   		UOWHF_Result[0].31:=0;
   		UOWHF_Result[1]:=UOWHF_Result[1] + 783475357+UOWHF_Add_c;
   		UOWHF_Add_c.1:=UOWHF_Result[1].31;
   		UOWHF_Result[1].31:=0;
   		UOWHF_Result[2]:=UOWHF_Result[2] + 293797280+UOWHF_Add_c;
   		UOWHF_Add_c.2:=UOWHF_Result[2].31;
   		UOWHF_Result[2].31:=0;
   		UOWHF_Result[3]:=UOWHF_Result[3] + 185650386+UOWHF_Add_c;
   		UOWHF_Add_c.3:=UOWHF_Result[3].31;
   		UOWHF_Result[3].31:=0;
   		UOWHF_Result[4]:=UOWHF_Result[4] + 976456778+UOWHF_Add_c;
   		UOWHF_Add_c.4:=UOWHF_Result[4].31;
   		UOWHF_Result[4].31:=0;
   		UOWHF_Result[5]:=UOWHF_Result[5] + 1830429797+UOWHF_Add_c;
   		UOWHF_Add_c.5:=UOWHF_Result[5].31;
   		UOWHF_Result[5].31:=0;
   		UOWHF_Result[6]:=UOWHF_Result[6] + 346921929+UOWHF_Add_c;
   		UOWHF_Add_c.6:=UOWHF_Result[6].31;
   		UOWHF_Result[6].31:=0;
   	End_If;
   	If UOWHF_Msg[1].[3] Then
   		UOWHF_Result[0]:=UOWHF_Result[0] + 542356735+UOWHF_Add_c;
   		UOWHF_Add_c.0:=UOWHF_Result[0].31;
   		UOWHF_Result[0].31:=0;
   		UOWHF_Result[1]:=UOWHF_Result[1] + 1471465957+UOWHF_Add_c;
   		UOWHF_Add_c.1:=UOWHF_Result[1].31;
   		UOWHF_Result[1].31:=0;
   		UOWHF_Result[2]:=UOWHF_Result[2] + 880885546+UOWHF_Add_c;
   		UOWHF_Add_c.2:=UOWHF_Result[2].31;
   		UOWHF_Result[2].31:=0;
   		UOWHF_Result[3]:=UOWHF_Result[3] + 1420715233+UOWHF_Add_c;
   		UOWHF_Add_c.3:=UOWHF_Result[3].31;
   		UOWHF_Result[3].31:=0;
   		UOWHF_Result[4]:=UOWHF_Result[4] + 974859291+UOWHF_Add_c;
   		UOWHF_Add_c.4:=UOWHF_Result[4].31;
   		UOWHF_Result[4].31:=0;
   		UOWHF_Result[5]:=UOWHF_Result[5] + 2135033399+UOWHF_Add_c;
   		UOWHF_Add_c.5:=UOWHF_Result[5].31;
   		UOWHF_Result[5].31:=0;
   		UOWHF_Result[6]:=UOWHF_Result[6] + 991907939+UOWHF_Add_c;
   		UOWHF_Add_c.6:=UOWHF_Result[6].31;
   		UOWHF_Result[6].31:=0;
   	End_If;
   	If UOWHF_Msg[1].[4] Then
   		UOWHF_Result[0]:=UOWHF_Result[0] + 233841843+UOWHF_Add_c;
   		UOWHF_Add_c.0:=UOWHF_Result[0].31;
   		UOWHF_Result[0].31:=0;
   		UOWHF_Result[1]:=UOWHF_Result[1] + 422275350+UOWHF_Add_c;
   		UOWHF_Add_c.1:=UOWHF_Result[1].31;
   		UOWHF_Result[1].31:=0;
   		UOWHF_Result[2]:=UOWHF_Result[2] + 758599260+UOWHF_Add_c;
   		UOWHF_Add_c.2:=UOWHF_Result[2].31;
   		UOWHF_Result[2].31:=0;
   		UOWHF_Result[3]:=UOWHF_Result[3] + 1065130774+UOWHF_Add_c;
   		UOWHF_Add_c.3:=UOWHF_Result[3].31;
   		UOWHF_Result[3].31:=0;
   		UOWHF_Result[4]:=UOWHF_Result[4] + 2001915225+UOWHF_Add_c;
   		UOWHF_Add_c.4:=UOWHF_Result[4].31;
   		UOWHF_Result[4].31:=0;
   		UOWHF_Result[5]:=UOWHF_Result[5] + 545495531+UOWHF_Add_c;
   		UOWHF_Add_c.5:=UOWHF_Result[5].31;
   		UOWHF_Result[5].31:=0;
   		UOWHF_Result[6]:=UOWHF_Result[6] + 296068018+UOWHF_Add_c;
   		UOWHF_Add_c.6:=UOWHF_Result[6].31;
   		UOWHF_Result[6].31:=0;
   	End_If;
   	If UOWHF_Msg[1].[5] Then
   		UOWHF_Result[0]:=UOWHF_Result[0] + 5724122+UOWHF_Add_c;
   		UOWHF_Add_c.0:=UOWHF_Result[0].31;
   		UOWHF_Result[0].31:=0;
   		UOWHF_Result[1]:=UOWHF_Result[1] + 218649241+UOWHF_Add_c;
   		UOWHF_Add_c.1:=UOWHF_Result[1].31;
   		UOWHF_Result[1].31:=0;
   		UOWHF_Result[2]:=UOWHF_Result[2] + 238121106+UOWHF_Add_c;
   		UOWHF_Add_c.2:=UOWHF_Result[2].31;
   		UOWHF_Result[2].31:=0;
   		UOWHF_Result[3]:=UOWHF_Result[3] + 729241869+UOWHF_Add_c;
   		UOWHF_Add_c.3:=UOWHF_Result[3].31;
   		UOWHF_Result[3].31:=0;
   		UOWHF_Result[4]:=UOWHF_Result[4] + 1651167024+UOWHF_Add_c;
   		UOWHF_Add_c.4:=UOWHF_Result[4].31;
   		UOWHF_Result[4].31:=0;
   		UOWHF_Result[5]:=UOWHF_Result[5] + 2110643339+UOWHF_Add_c;
   		UOWHF_Add_c.5:=UOWHF_Result[5].31;
   		UOWHF_Result[5].31:=0;
   		UOWHF_Result[6]:=UOWHF_Result[6] + 1917524854+UOWHF_Add_c;
   		UOWHF_Add_c.6:=UOWHF_Result[6].31;
   		UOWHF_Result[6].31:=0;
   	End_If;
   	If UOWHF_Msg[1].[6] Then
   		UOWHF_Result[0]:=UOWHF_Result[0] + 573579892+UOWHF_Add_c;
   		UOWHF_Add_c.0:=UOWHF_Result[0].31;
   		UOWHF_Result[0].31:=0;
   		UOWHF_Result[1]:=UOWHF_Result[1] + 1647169020+UOWHF_Add_c;
   		UOWHF_Add_c.1:=UOWHF_Result[1].31;
   		UOWHF_Result[1].31:=0;
   		UOWHF_Result[2]:=UOWHF_Result[2] + 144695872+UOWHF_Add_c;
   		UOWHF_Add_c.2:=UOWHF_Result[2].31;
   		UOWHF_Result[2].31:=0;
   		UOWHF_Result[3]:=UOWHF_Result[3] + 858449959+UOWHF_Add_c;
   		UOWHF_Add_c.3:=UOWHF_Result[3].31;
   		UOWHF_Result[3].31:=0;
   		UOWHF_Result[4]:=UOWHF_Result[4] + 514618441+UOWHF_Add_c;
   		UOWHF_Add_c.4:=UOWHF_Result[4].31;
   		UOWHF_Result[4].31:=0;
   		UOWHF_Result[5]:=UOWHF_Result[5] + 38664886+UOWHF_Add_c;
   		UOWHF_Add_c.5:=UOWHF_Result[5].31;
   		UOWHF_Result[5].31:=0;
   		UOWHF_Result[6]:=UOWHF_Result[6] + 2115485271+UOWHF_Add_c;
   		UOWHF_Add_c.6:=UOWHF_Result[6].31;
   		UOWHF_Result[6].31:=0;
   	End_If;
   	If UOWHF_Msg[1].[7] Then
   		UOWHF_Result[0]:=UOWHF_Result[0] + 1170004469+UOWHF_Add_c;
   		UOWHF_Add_c.0:=UOWHF_Result[0].31;
   		UOWHF_Result[0].31:=0;
   		UOWHF_Result[1]:=UOWHF_Result[1] + 37314947+UOWHF_Add_c;
   		UOWHF_Add_c.1:=UOWHF_Result[1].31;
   		UOWHF_Result[1].31:=0;
   		UOWHF_Result[2]:=UOWHF_Result[2] + 946474451+UOWHF_Add_c;
   		UOWHF_Add_c.2:=UOWHF_Result[2].31;
   		UOWHF_Result[2].31:=0;
   		UOWHF_Result[3]:=UOWHF_Result[3] + 896038805+UOWHF_Add_c;
   		UOWHF_Add_c.3:=UOWHF_Result[3].31;
   		UOWHF_Result[3].31:=0;
   		UOWHF_Result[4]:=UOWHF_Result[4] + 2098536983+UOWHF_Add_c;
   		UOWHF_Add_c.4:=UOWHF_Result[4].31;
   		UOWHF_Result[4].31:=0;
   		UOWHF_Result[5]:=UOWHF_Result[5] + 1225593261+UOWHF_Add_c;
   		UOWHF_Add_c.5:=UOWHF_Result[5].31;
   		UOWHF_Result[5].31:=0;
   		UOWHF_Result[6]:=UOWHF_Result[6] + 1353408681+UOWHF_Add_c;
   		UOWHF_Add_c.6:=UOWHF_Result[6].31;
   		UOWHF_Result[6].31:=0;
   	End_If;
   	If UOWHF_Msg[1].[8] Then
   		UOWHF_Result[0]:=UOWHF_Result[0] + 1872283162+UOWHF_Add_c;
   		UOWHF_Add_c.0:=UOWHF_Result[0].31;
   		UOWHF_Result[0].31:=0;
   		UOWHF_Result[1]:=UOWHF_Result[1] + 1856697315+UOWHF_Add_c;
   		UOWHF_Add_c.1:=UOWHF_Result[1].31;
   		UOWHF_Result[1].31:=0;
   		UOWHF_Result[2]:=UOWHF_Result[2] + 360372569+UOWHF_Add_c;
   		UOWHF_Add_c.2:=UOWHF_Result[2].31;
   		UOWHF_Result[2].31:=0;
   		UOWHF_Result[3]:=UOWHF_Result[3] + 726928957+UOWHF_Add_c;
   		UOWHF_Add_c.3:=UOWHF_Result[3].31;
   		UOWHF_Result[3].31:=0;
   		UOWHF_Result[4]:=UOWHF_Result[4] + 159244533+UOWHF_Add_c;
   		UOWHF_Add_c.4:=UOWHF_Result[4].31;
   		UOWHF_Result[4].31:=0;
   		UOWHF_Result[5]:=UOWHF_Result[5] + 218947815+UOWHF_Add_c;
   		UOWHF_Add_c.5:=UOWHF_Result[5].31;
   		UOWHF_Result[5].31:=0;
   		UOWHF_Result[6]:=UOWHF_Result[6] + 1781099399+UOWHF_Add_c;
   		UOWHF_Add_c.6:=UOWHF_Result[6].31;
   		UOWHF_Result[6].31:=0;
   	End_If;
   	If UOWHF_Msg[1].[9] Then
   		UOWHF_Result[0]:=UOWHF_Result[0] + 1141680914+UOWHF_Add_c;
   		UOWHF_Add_c.0:=UOWHF_Result[0].31;
   		UOWHF_Result[0].31:=0;
   		UOWHF_Result[1]:=UOWHF_Result[1] + 501780076+UOWHF_Add_c;
   		UOWHF_Add_c.1:=UOWHF_Result[1].31;
   		UOWHF_Result[1].31:=0;
   		UOWHF_Result[2]:=UOWHF_Result[2] + 1857845686+UOWHF_Add_c;
   		UOWHF_Add_c.2:=UOWHF_Result[2].31;
   		UOWHF_Result[2].31:=0;
   		UOWHF_Result[3]:=UOWHF_Result[3] + 1524263353+UOWHF_Add_c;
   		UOWHF_Add_c.3:=UOWHF_Result[3].31;
   		UOWHF_Result[3].31:=0;
   		UOWHF_Result[4]:=UOWHF_Result[4] + 337597395+UOWHF_Add_c;
   		UOWHF_Add_c.4:=UOWHF_Result[4].31;
   		UOWHF_Result[4].31:=0;
   		UOWHF_Result[5]:=UOWHF_Result[5] + 479430851+UOWHF_Add_c;
   		UOWHF_Add_c.5:=UOWHF_Result[5].31;
   		UOWHF_Result[5].31:=0;
   		UOWHF_Result[6]:=UOWHF_Result[6] + 1673187600+UOWHF_Add_c;
   		UOWHF_Add_c.6:=UOWHF_Result[6].31;
   		UOWHF_Result[6].31:=0;
   	End_If;
   	If UOWHF_Msg[1].[10] Then
   		UOWHF_Result[0]:=UOWHF_Result[0] + 242125945+UOWHF_Add_c;
   		UOWHF_Add_c.0:=UOWHF_Result[0].31;
   		UOWHF_Result[0].31:=0;
   		UOWHF_Result[1]:=UOWHF_Result[1] + 640016629+UOWHF_Add_c;
   		UOWHF_Add_c.1:=UOWHF_Result[1].31;
   		UOWHF_Result[1].31:=0;
   		UOWHF_Result[2]:=UOWHF_Result[2] + 2080248052+UOWHF_Add_c;
   		UOWHF_Add_c.2:=UOWHF_Result[2].31;
   		UOWHF_Result[2].31:=0;
   		UOWHF_Result[3]:=UOWHF_Result[3] + 1952927158+UOWHF_Add_c;
   		UOWHF_Add_c.3:=UOWHF_Result[3].31;
   		UOWHF_Result[3].31:=0;
   		UOWHF_Result[4]:=UOWHF_Result[4] + 1703045187+UOWHF_Add_c;
   		UOWHF_Add_c.4:=UOWHF_Result[4].31;
   		UOWHF_Result[4].31:=0;
   		UOWHF_Result[5]:=UOWHF_Result[5] + 1628740462+UOWHF_Add_c;
   		UOWHF_Add_c.5:=UOWHF_Result[5].31;
   		UOWHF_Result[5].31:=0;
   		UOWHF_Result[6]:=UOWHF_Result[6] + 546275254+UOWHF_Add_c;
   		UOWHF_Add_c.6:=UOWHF_Result[6].31;
   		UOWHF_Result[6].31:=0;
   	End_If;
   	If UOWHF_Msg[1].[11] Then
   		UOWHF_Result[0]:=UOWHF_Result[0] + 1214351459+UOWHF_Add_c;
   		UOWHF_Add_c.0:=UOWHF_Result[0].31;
   		UOWHF_Result[0].31:=0;
   		UOWHF_Result[1]:=UOWHF_Result[1] + 1585902034+UOWHF_Add_c;
   		UOWHF_Add_c.1:=UOWHF_Result[1].31;
   		UOWHF_Result[1].31:=0;
   		UOWHF_Result[2]:=UOWHF_Result[2] + 2020777692+UOWHF_Add_c;
   		UOWHF_Add_c.2:=UOWHF_Result[2].31;
   		UOWHF_Result[2].31:=0;
   		UOWHF_Result[3]:=UOWHF_Result[3] + 831190818+UOWHF_Add_c;
   		UOWHF_Add_c.3:=UOWHF_Result[3].31;
   		UOWHF_Result[3].31:=0;
   		UOWHF_Result[4]:=UOWHF_Result[4] + 1956522628+UOWHF_Add_c;
   		UOWHF_Add_c.4:=UOWHF_Result[4].31;
   		UOWHF_Result[4].31:=0;
   		UOWHF_Result[5]:=UOWHF_Result[5] + 1924488146+UOWHF_Add_c;
   		UOWHF_Add_c.5:=UOWHF_Result[5].31;
   		UOWHF_Result[5].31:=0;
   		UOWHF_Result[6]:=UOWHF_Result[6] + 1582768083+UOWHF_Add_c;
   		UOWHF_Add_c.6:=UOWHF_Result[6].31;
   		UOWHF_Result[6].31:=0;
   	End_If;
   	If UOWHF_Msg[1].[12] Then
   		UOWHF_Result[0]:=UOWHF_Result[0] + 1902205147+UOWHF_Add_c;
   		UOWHF_Add_c.0:=UOWHF_Result[0].31;
   		UOWHF_Result[0].31:=0;
   		UOWHF_Result[1]:=UOWHF_Result[1] + 1414042614+UOWHF_Add_c;
   		UOWHF_Add_c.1:=UOWHF_Result[1].31;
   		UOWHF_Result[1].31:=0;
   		UOWHF_Result[2]:=UOWHF_Result[2] + 1252562892+UOWHF_Add_c;
   		UOWHF_Add_c.2:=UOWHF_Result[2].31;
   		UOWHF_Result[2].31:=0;
   		UOWHF_Result[3]:=UOWHF_Result[3] + 1986955796+UOWHF_Add_c;
   		UOWHF_Add_c.3:=UOWHF_Result[3].31;
   		UOWHF_Result[3].31:=0;
   		UOWHF_Result[4]:=UOWHF_Result[4] + 1280256904+UOWHF_Add_c;
   		UOWHF_Add_c.4:=UOWHF_Result[4].31;
   		UOWHF_Result[4].31:=0;
   		UOWHF_Result[5]:=UOWHF_Result[5] + 1879967415+UOWHF_Add_c;
   		UOWHF_Add_c.5:=UOWHF_Result[5].31;
   		UOWHF_Result[5].31:=0;
   		UOWHF_Result[6]:=UOWHF_Result[6] + 2127199076+UOWHF_Add_c;
   		UOWHF_Add_c.6:=UOWHF_Result[6].31;
   		UOWHF_Result[6].31:=0;
   	End_If;
   	If UOWHF_Msg[1].[13] Then
   		UOWHF_Result[0]:=UOWHF_Result[0] + 308710562+UOWHF_Add_c;
   		UOWHF_Add_c.0:=UOWHF_Result[0].31;
   		UOWHF_Result[0].31:=0;
   		UOWHF_Result[1]:=UOWHF_Result[1] + 840066539+UOWHF_Add_c;
   		UOWHF_Add_c.1:=UOWHF_Result[1].31;
   		UOWHF_Result[1].31:=0;
   		UOWHF_Result[2]:=UOWHF_Result[2] + 2112096411+UOWHF_Add_c;
   		UOWHF_Add_c.2:=UOWHF_Result[2].31;
   		UOWHF_Result[2].31:=0;
   		UOWHF_Result[3]:=UOWHF_Result[3] + 430276806+UOWHF_Add_c;
   		UOWHF_Add_c.3:=UOWHF_Result[3].31;
   		UOWHF_Result[3].31:=0;
   		UOWHF_Result[4]:=UOWHF_Result[4] + 1656622260+UOWHF_Add_c;
   		UOWHF_Add_c.4:=UOWHF_Result[4].31;
   		UOWHF_Result[4].31:=0;
   		UOWHF_Result[5]:=UOWHF_Result[5] + 1475134647+UOWHF_Add_c;
   		UOWHF_Add_c.5:=UOWHF_Result[5].31;
   		UOWHF_Result[5].31:=0;
   		UOWHF_Result[6]:=UOWHF_Result[6] + 1218741234+UOWHF_Add_c;
   		UOWHF_Add_c.6:=UOWHF_Result[6].31;
   		UOWHF_Result[6].31:=0;
   	End_If;
   	If UOWHF_Msg[1].[14] Then
   		UOWHF_Result[0]:=UOWHF_Result[0] + 79982991+UOWHF_Add_c;
   		UOWHF_Add_c.0:=UOWHF_Result[0].31;
   		UOWHF_Result[0].31:=0;
   		UOWHF_Result[1]:=UOWHF_Result[1] + 1048582461+UOWHF_Add_c;
   		UOWHF_Add_c.1:=UOWHF_Result[1].31;
   		UOWHF_Result[1].31:=0;
   		UOWHF_Result[2]:=UOWHF_Result[2] + 1041482528+UOWHF_Add_c;
   		UOWHF_Add_c.2:=UOWHF_Result[2].31;
   		UOWHF_Result[2].31:=0;
   		UOWHF_Result[3]:=UOWHF_Result[3] + 1202571175+UOWHF_Add_c;
   		UOWHF_Add_c.3:=UOWHF_Result[3].31;
   		UOWHF_Result[3].31:=0;
   		UOWHF_Result[4]:=UOWHF_Result[4] + 429088756+UOWHF_Add_c;
   		UOWHF_Add_c.4:=UOWHF_Result[4].31;
   		UOWHF_Result[4].31:=0;
   		UOWHF_Result[5]:=UOWHF_Result[5] + 1706637211+UOWHF_Add_c;
   		UOWHF_Add_c.5:=UOWHF_Result[5].31;
   		UOWHF_Result[5].31:=0;
   		UOWHF_Result[6]:=UOWHF_Result[6] + 1523304685+UOWHF_Add_c;
   		UOWHF_Add_c.6:=UOWHF_Result[6].31;
   		UOWHF_Result[6].31:=0;
   	End_If;
   	If UOWHF_Msg[1].[15] Then
   		UOWHF_Result[0]:=UOWHF_Result[0] + 1151565721+UOWHF_Add_c;
   		UOWHF_Add_c.0:=UOWHF_Result[0].31;
   		UOWHF_Result[0].31:=0;
   		UOWHF_Result[1]:=UOWHF_Result[1] + 326738685+UOWHF_Add_c;
   		UOWHF_Add_c.1:=UOWHF_Result[1].31;
   		UOWHF_Result[1].31:=0;
   		UOWHF_Result[2]:=UOWHF_Result[2] + 848077496+UOWHF_Add_c;
   		UOWHF_Add_c.2:=UOWHF_Result[2].31;
   		UOWHF_Result[2].31:=0;
   		UOWHF_Result[3]:=UOWHF_Result[3] + 1977621819+UOWHF_Add_c;
   		UOWHF_Add_c.3:=UOWHF_Result[3].31;
   		UOWHF_Result[3].31:=0;
   		UOWHF_Result[4]:=UOWHF_Result[4] + 8183745+UOWHF_Add_c;
   		UOWHF_Add_c.4:=UOWHF_Result[4].31;
   		UOWHF_Result[4].31:=0;
   		UOWHF_Result[5]:=UOWHF_Result[5] + 1696313996+UOWHF_Add_c;
   		UOWHF_Add_c.5:=UOWHF_Result[5].31;
   		UOWHF_Result[5].31:=0;
   		UOWHF_Result[6]:=UOWHF_Result[6] + 2057304671+UOWHF_Add_c;
   		UOWHF_Add_c.6:=UOWHF_Result[6].31;
   		UOWHF_Result[6].31:=0;
   	End_If;
   	If UOWHF_Msg[1].[16] Then
   		UOWHF_Result[0]:=UOWHF_Result[0] + 374952423+UOWHF_Add_c;
   		UOWHF_Add_c.0:=UOWHF_Result[0].31;
   		UOWHF_Result[0].31:=0;
   		UOWHF_Result[1]:=UOWHF_Result[1] + 1823443600+UOWHF_Add_c;
   		UOWHF_Add_c.1:=UOWHF_Result[1].31;
   		UOWHF_Result[1].31:=0;
   		UOWHF_Result[2]:=UOWHF_Result[2] + 1962739745+UOWHF_Add_c;
   		UOWHF_Add_c.2:=UOWHF_Result[2].31;
   		UOWHF_Result[2].31:=0;
   		UOWHF_Result[3]:=UOWHF_Result[3] + 494646021+UOWHF_Add_c;
   		UOWHF_Add_c.3:=UOWHF_Result[3].31;
   		UOWHF_Result[3].31:=0;
   		UOWHF_Result[4]:=UOWHF_Result[4] + 2102427342+UOWHF_Add_c;
   		UOWHF_Add_c.4:=UOWHF_Result[4].31;
   		UOWHF_Result[4].31:=0;
   		UOWHF_Result[5]:=UOWHF_Result[5] + 1782471367+UOWHF_Add_c;
   		UOWHF_Add_c.5:=UOWHF_Result[5].31;
   		UOWHF_Result[5].31:=0;
   		UOWHF_Result[6]:=UOWHF_Result[6] + 861507114+UOWHF_Add_c;
   		UOWHF_Add_c.6:=UOWHF_Result[6].31;
   		UOWHF_Result[6].31:=0;
   	End_If;
   	If UOWHF_Msg[1].[17] Then
   		UOWHF_Result[0]:=UOWHF_Result[0] + 432199441+UOWHF_Add_c;
   		UOWHF_Add_c.0:=UOWHF_Result[0].31;
   		UOWHF_Result[0].31:=0;
   		UOWHF_Result[1]:=UOWHF_Result[1] + 828673085+UOWHF_Add_c;
   		UOWHF_Add_c.1:=UOWHF_Result[1].31;
   		UOWHF_Result[1].31:=0;
   		UOWHF_Result[2]:=UOWHF_Result[2] + 1984216486+UOWHF_Add_c;
   		UOWHF_Add_c.2:=UOWHF_Result[2].31;
   		UOWHF_Result[2].31:=0;
   		UOWHF_Result[3]:=UOWHF_Result[3] + 1064724900+UOWHF_Add_c;
   		UOWHF_Add_c.3:=UOWHF_Result[3].31;
   		UOWHF_Result[3].31:=0;
   		UOWHF_Result[4]:=UOWHF_Result[4] + 874774630+UOWHF_Add_c;
   		UOWHF_Add_c.4:=UOWHF_Result[4].31;
   		UOWHF_Result[4].31:=0;
   		UOWHF_Result[5]:=UOWHF_Result[5] + 21515165+UOWHF_Add_c;
   		UOWHF_Add_c.5:=UOWHF_Result[5].31;
   		UOWHF_Result[5].31:=0;
   		UOWHF_Result[6]:=UOWHF_Result[6] + 1481985786+UOWHF_Add_c;
   		UOWHF_Add_c.6:=UOWHF_Result[6].31;
   		UOWHF_Result[6].31:=0;
   	End_If;
   	If UOWHF_Msg[1].[18] Then
   		UOWHF_Result[0]:=UOWHF_Result[0] + 1771683016+UOWHF_Add_c;
   		UOWHF_Add_c.0:=UOWHF_Result[0].31;
   		UOWHF_Result[0].31:=0;
   		UOWHF_Result[1]:=UOWHF_Result[1] + 1893376172+UOWHF_Add_c;
   		UOWHF_Add_c.1:=UOWHF_Result[1].31;
   		UOWHF_Result[1].31:=0;
   		UOWHF_Result[2]:=UOWHF_Result[2] + 589589901+UOWHF_Add_c;
   		UOWHF_Add_c.2:=UOWHF_Result[2].31;
   		UOWHF_Result[2].31:=0;
   		UOWHF_Result[3]:=UOWHF_Result[3] + 1014880440+UOWHF_Add_c;
   		UOWHF_Add_c.3:=UOWHF_Result[3].31;
   		UOWHF_Result[3].31:=0;
   		UOWHF_Result[4]:=UOWHF_Result[4] + 1125259377+UOWHF_Add_c;
   		UOWHF_Add_c.4:=UOWHF_Result[4].31;
   		UOWHF_Result[4].31:=0;
   		UOWHF_Result[5]:=UOWHF_Result[5] + 1266464258+UOWHF_Add_c;
   		UOWHF_Add_c.5:=UOWHF_Result[5].31;
   		UOWHF_Result[5].31:=0;
   		UOWHF_Result[6]:=UOWHF_Result[6] + 2138531095+UOWHF_Add_c;
   		UOWHF_Add_c.6:=UOWHF_Result[6].31;
   		UOWHF_Result[6].31:=0;
   	End_If;
   	If UOWHF_Msg[1].[19] Then
   		UOWHF_Result[0]:=UOWHF_Result[0] + 702390516+UOWHF_Add_c;
   		UOWHF_Add_c.0:=UOWHF_Result[0].31;
   		UOWHF_Result[0].31:=0;
   		UOWHF_Result[1]:=UOWHF_Result[1] + 1522466915+UOWHF_Add_c;
   		UOWHF_Add_c.1:=UOWHF_Result[1].31;
   		UOWHF_Result[1].31:=0;
   		UOWHF_Result[2]:=UOWHF_Result[2] + 143129679+UOWHF_Add_c;
   		UOWHF_Add_c.2:=UOWHF_Result[2].31;
   		UOWHF_Result[2].31:=0;
   		UOWHF_Result[3]:=UOWHF_Result[3] + 666937844+UOWHF_Add_c;
   		UOWHF_Add_c.3:=UOWHF_Result[3].31;
   		UOWHF_Result[3].31:=0;
   		UOWHF_Result[4]:=UOWHF_Result[4] + 1262542875+UOWHF_Add_c;
   		UOWHF_Add_c.4:=UOWHF_Result[4].31;
   		UOWHF_Result[4].31:=0;
   		UOWHF_Result[5]:=UOWHF_Result[5] + 1076685305+UOWHF_Add_c;
   		UOWHF_Add_c.5:=UOWHF_Result[5].31;
   		UOWHF_Result[5].31:=0;
   		UOWHF_Result[6]:=UOWHF_Result[6] + 494452534+UOWHF_Add_c;
   		UOWHF_Add_c.6:=UOWHF_Result[6].31;
   		UOWHF_Result[6].31:=0;
   	End_If;
   	If UOWHF_Msg[1].[20] Then
   		UOWHF_Result[0]:=UOWHF_Result[0] + 1156353219+UOWHF_Add_c;
   		UOWHF_Add_c.0:=UOWHF_Result[0].31;
   		UOWHF_Result[0].31:=0;
   		UOWHF_Result[1]:=UOWHF_Result[1] + 1843399297+UOWHF_Add_c;
   		UOWHF_Add_c.1:=UOWHF_Result[1].31;
   		UOWHF_Result[1].31:=0;
   		UOWHF_Result[2]:=UOWHF_Result[2] + 777057182+UOWHF_Add_c;
   		UOWHF_Add_c.2:=UOWHF_Result[2].31;
   		UOWHF_Result[2].31:=0;
   		UOWHF_Result[3]:=UOWHF_Result[3] + 933746277+UOWHF_Add_c;
   		UOWHF_Add_c.3:=UOWHF_Result[3].31;
   		UOWHF_Result[3].31:=0;
   		UOWHF_Result[4]:=UOWHF_Result[4] + 1158149847+UOWHF_Add_c;
   		UOWHF_Add_c.4:=UOWHF_Result[4].31;
   		UOWHF_Result[4].31:=0;
   		UOWHF_Result[5]:=UOWHF_Result[5] + 653472915+UOWHF_Add_c;
   		UOWHF_Add_c.5:=UOWHF_Result[5].31;
   		UOWHF_Result[5].31:=0;
   		UOWHF_Result[6]:=UOWHF_Result[6] + 1413034676+UOWHF_Add_c;
   		UOWHF_Add_c.6:=UOWHF_Result[6].31;
   		UOWHF_Result[6].31:=0;
   	End_If;
   	If UOWHF_Msg[1].[21] Then
   		UOWHF_Result[0]:=UOWHF_Result[0] + 1572421213+UOWHF_Add_c;
   		UOWHF_Add_c.0:=UOWHF_Result[0].31;
   		UOWHF_Result[0].31:=0;
   		UOWHF_Result[1]:=UOWHF_Result[1] + 88389224+UOWHF_Add_c;
   		UOWHF_Add_c.1:=UOWHF_Result[1].31;
   		UOWHF_Result[1].31:=0;
   		UOWHF_Result[2]:=UOWHF_Result[2] + 400840719+UOWHF_Add_c;
   		UOWHF_Add_c.2:=UOWHF_Result[2].31;
   		UOWHF_Result[2].31:=0;
   		UOWHF_Result[3]:=UOWHF_Result[3] + 77634928+UOWHF_Add_c;
   		UOWHF_Add_c.3:=UOWHF_Result[3].31;
   		UOWHF_Result[3].31:=0;
   		UOWHF_Result[4]:=UOWHF_Result[4] + 930991932+UOWHF_Add_c;
   		UOWHF_Add_c.4:=UOWHF_Result[4].31;
   		UOWHF_Result[4].31:=0;
   		UOWHF_Result[5]:=UOWHF_Result[5] + 728144988+UOWHF_Add_c;
   		UOWHF_Add_c.5:=UOWHF_Result[5].31;
   		UOWHF_Result[5].31:=0;
   		UOWHF_Result[6]:=UOWHF_Result[6] + 615317385+UOWHF_Add_c;
   		UOWHF_Add_c.6:=UOWHF_Result[6].31;
   		UOWHF_Result[6].31:=0;
   	End_If;
   	If UOWHF_Msg[1].[22] Then
   		UOWHF_Result[0]:=UOWHF_Result[0] + 621466345+UOWHF_Add_c;
   		UOWHF_Add_c.0:=UOWHF_Result[0].31;
   		UOWHF_Result[0].31:=0;
   		UOWHF_Result[1]:=UOWHF_Result[1] + 1585265844+UOWHF_Add_c;
   		UOWHF_Add_c.1:=UOWHF_Result[1].31;
   		UOWHF_Result[1].31:=0;
   		UOWHF_Result[2]:=UOWHF_Result[2] + 329909774+UOWHF_Add_c;
   		UOWHF_Add_c.2:=UOWHF_Result[2].31;
   		UOWHF_Result[2].31:=0;
   		UOWHF_Result[3]:=UOWHF_Result[3] + 1704616883+UOWHF_Add_c;
   		UOWHF_Add_c.3:=UOWHF_Result[3].31;
   		UOWHF_Result[3].31:=0;
   		UOWHF_Result[4]:=UOWHF_Result[4] + 887994120+UOWHF_Add_c;
   		UOWHF_Add_c.4:=UOWHF_Result[4].31;
   		UOWHF_Result[4].31:=0;
   		UOWHF_Result[5]:=UOWHF_Result[5] + 2033117695+UOWHF_Add_c;
   		UOWHF_Add_c.5:=UOWHF_Result[5].31;
   		UOWHF_Result[5].31:=0;
   		UOWHF_Result[6]:=UOWHF_Result[6] + 1261571647+UOWHF_Add_c;
   		UOWHF_Add_c.6:=UOWHF_Result[6].31;
   		UOWHF_Result[6].31:=0;
   	End_If;
   	If UOWHF_Msg[1].[23] Then
   		UOWHF_Result[0]:=UOWHF_Result[0] + 1919220287+UOWHF_Add_c;
   		UOWHF_Add_c.0:=UOWHF_Result[0].31;
   		UOWHF_Result[0].31:=0;
   		UOWHF_Result[1]:=UOWHF_Result[1] + 1329200192+UOWHF_Add_c;
   		UOWHF_Add_c.1:=UOWHF_Result[1].31;
   		UOWHF_Result[1].31:=0;
   		UOWHF_Result[2]:=UOWHF_Result[2] + 2036885514+UOWHF_Add_c;
   		UOWHF_Add_c.2:=UOWHF_Result[2].31;
   		UOWHF_Result[2].31:=0;
   		UOWHF_Result[3]:=UOWHF_Result[3] + 1069469832+UOWHF_Add_c;
   		UOWHF_Add_c.3:=UOWHF_Result[3].31;
   		UOWHF_Result[3].31:=0;
   		UOWHF_Result[4]:=UOWHF_Result[4] + 736892868+UOWHF_Add_c;
   		UOWHF_Add_c.4:=UOWHF_Result[4].31;
   		UOWHF_Result[4].31:=0;
   		UOWHF_Result[5]:=UOWHF_Result[5] + 1241914734+UOWHF_Add_c;
   		UOWHF_Add_c.5:=UOWHF_Result[5].31;
   		UOWHF_Result[5].31:=0;
   		UOWHF_Result[6]:=UOWHF_Result[6] + 853099692+UOWHF_Add_c;
   		UOWHF_Add_c.6:=UOWHF_Result[6].31;
   		UOWHF_Result[6].31:=0;
   	End_If;
   	If UOWHF_Msg[1].[24] Then
   		UOWHF_Result[0]:=UOWHF_Result[0] + 997973851+UOWHF_Add_c;
   		UOWHF_Add_c.0:=UOWHF_Result[0].31;
   		UOWHF_Result[0].31:=0;
   		UOWHF_Result[1]:=UOWHF_Result[1] + 744436970+UOWHF_Add_c;
   		UOWHF_Add_c.1:=UOWHF_Result[1].31;
   		UOWHF_Result[1].31:=0;
   		UOWHF_Result[2]:=UOWHF_Result[2] + 2040904751+UOWHF_Add_c;
   		UOWHF_Add_c.2:=UOWHF_Result[2].31;
   		UOWHF_Result[2].31:=0;
   		UOWHF_Result[3]:=UOWHF_Result[3] + 877190201+UOWHF_Add_c;
   		UOWHF_Add_c.3:=UOWHF_Result[3].31;
   		UOWHF_Result[3].31:=0;
   		UOWHF_Result[4]:=UOWHF_Result[4] + 1629723595+UOWHF_Add_c;
   		UOWHF_Add_c.4:=UOWHF_Result[4].31;
   		UOWHF_Result[4].31:=0;
   		UOWHF_Result[5]:=UOWHF_Result[5] + 1324262795+UOWHF_Add_c;
   		UOWHF_Add_c.5:=UOWHF_Result[5].31;
   		UOWHF_Result[5].31:=0;
   		UOWHF_Result[6]:=UOWHF_Result[6] + 455895855+UOWHF_Add_c;
   		UOWHF_Add_c.6:=UOWHF_Result[6].31;
   		UOWHF_Result[6].31:=0;
   	End_If;
   	If UOWHF_Msg[1].[25] Then
   		UOWHF_Result[0]:=UOWHF_Result[0] + 1233884413+UOWHF_Add_c;
   		UOWHF_Add_c.0:=UOWHF_Result[0].31;
   		UOWHF_Result[0].31:=0;
   		UOWHF_Result[1]:=UOWHF_Result[1] + 1172639779+UOWHF_Add_c;
   		UOWHF_Add_c.1:=UOWHF_Result[1].31;
   		UOWHF_Result[1].31:=0;
   		UOWHF_Result[2]:=UOWHF_Result[2] + 1187965169+UOWHF_Add_c;
   		UOWHF_Add_c.2:=UOWHF_Result[2].31;
   		UOWHF_Result[2].31:=0;
   		UOWHF_Result[3]:=UOWHF_Result[3] + 1965583593+UOWHF_Add_c;
   		UOWHF_Add_c.3:=UOWHF_Result[3].31;
   		UOWHF_Result[3].31:=0;
   		UOWHF_Result[4]:=UOWHF_Result[4] + 148415583+UOWHF_Add_c;
   		UOWHF_Add_c.4:=UOWHF_Result[4].31;
   		UOWHF_Result[4].31:=0;
   		UOWHF_Result[5]:=UOWHF_Result[5] + 1681123673+UOWHF_Add_c;
   		UOWHF_Add_c.5:=UOWHF_Result[5].31;
   		UOWHF_Result[5].31:=0;
   		UOWHF_Result[6]:=UOWHF_Result[6] + 231213872+UOWHF_Add_c;
   		UOWHF_Add_c.6:=UOWHF_Result[6].31;
   		UOWHF_Result[6].31:=0;
   	End_If;
   	If UOWHF_Msg[1].[26] Then
   		UOWHF_Result[0]:=UOWHF_Result[0] + 1384429274+UOWHF_Add_c;
   		UOWHF_Add_c.0:=UOWHF_Result[0].31;
   		UOWHF_Result[0].31:=0;
   		UOWHF_Result[1]:=UOWHF_Result[1] + 1404381353+UOWHF_Add_c;
   		UOWHF_Add_c.1:=UOWHF_Result[1].31;
   		UOWHF_Result[1].31:=0;
   		UOWHF_Result[2]:=UOWHF_Result[2] + 604171081+UOWHF_Add_c;
   		UOWHF_Add_c.2:=UOWHF_Result[2].31;
   		UOWHF_Result[2].31:=0;
   		UOWHF_Result[3]:=UOWHF_Result[3] + 989237533+UOWHF_Add_c;
   		UOWHF_Add_c.3:=UOWHF_Result[3].31;
   		UOWHF_Result[3].31:=0;
   		UOWHF_Result[4]:=UOWHF_Result[4] + 1309759137+UOWHF_Add_c;
   		UOWHF_Add_c.4:=UOWHF_Result[4].31;
   		UOWHF_Result[4].31:=0;
   		UOWHF_Result[5]:=UOWHF_Result[5] + 678109269+UOWHF_Add_c;
   		UOWHF_Add_c.5:=UOWHF_Result[5].31;
   		UOWHF_Result[5].31:=0;
   		UOWHF_Result[6]:=UOWHF_Result[6] + 1506438700+UOWHF_Add_c;
   		UOWHF_Add_c.6:=UOWHF_Result[6].31;
   		UOWHF_Result[6].31:=0;
   	End_If;
   	If UOWHF_Msg[1].[27] Then
   		UOWHF_Result[0]:=UOWHF_Result[0] + 1630240536+UOWHF_Add_c;
   		UOWHF_Add_c.0:=UOWHF_Result[0].31;
   		UOWHF_Result[0].31:=0;
   		UOWHF_Result[1]:=UOWHF_Result[1] + 1425405810+UOWHF_Add_c;
   		UOWHF_Add_c.1:=UOWHF_Result[1].31;
   		UOWHF_Result[1].31:=0;
   		UOWHF_Result[2]:=UOWHF_Result[2] + 2087621973+UOWHF_Add_c;
   		UOWHF_Add_c.2:=UOWHF_Result[2].31;
   		UOWHF_Result[2].31:=0;
   		UOWHF_Result[3]:=UOWHF_Result[3] + 1431955454+UOWHF_Add_c;
   		UOWHF_Add_c.3:=UOWHF_Result[3].31;
   		UOWHF_Result[3].31:=0;
   		UOWHF_Result[4]:=UOWHF_Result[4] + 1211813660+UOWHF_Add_c;
   		UOWHF_Add_c.4:=UOWHF_Result[4].31;
   		UOWHF_Result[4].31:=0;
   		UOWHF_Result[5]:=UOWHF_Result[5] + 44221546+UOWHF_Add_c;
   		UOWHF_Add_c.5:=UOWHF_Result[5].31;
   		UOWHF_Result[5].31:=0;
   		UOWHF_Result[6]:=UOWHF_Result[6] + 1700714287+UOWHF_Add_c;
   		UOWHF_Add_c.6:=UOWHF_Result[6].31;
   		UOWHF_Result[6].31:=0;
   	End_If;
   	If UOWHF_Msg[1].[28] Then
   		UOWHF_Result[0]:=UOWHF_Result[0] + 2018244125+UOWHF_Add_c;
   		UOWHF_Add_c.0:=UOWHF_Result[0].31;
   		UOWHF_Result[0].31:=0;
   		UOWHF_Result[1]:=UOWHF_Result[1] + 529957975+UOWHF_Add_c;
   		UOWHF_Add_c.1:=UOWHF_Result[1].31;
   		UOWHF_Result[1].31:=0;
   		UOWHF_Result[2]:=UOWHF_Result[2] + 691952083+UOWHF_Add_c;
   		UOWHF_Add_c.2:=UOWHF_Result[2].31;
   		UOWHF_Result[2].31:=0;
   		UOWHF_Result[3]:=UOWHF_Result[3] + 405329013+UOWHF_Add_c;
   		UOWHF_Add_c.3:=UOWHF_Result[3].31;
   		UOWHF_Result[3].31:=0;
   		UOWHF_Result[4]:=UOWHF_Result[4] + 1980445743+UOWHF_Add_c;
   		UOWHF_Add_c.4:=UOWHF_Result[4].31;
   		UOWHF_Result[4].31:=0;
   		UOWHF_Result[5]:=UOWHF_Result[5] + 1515594315+UOWHF_Add_c;
   		UOWHF_Add_c.5:=UOWHF_Result[5].31;
   		UOWHF_Result[5].31:=0;
   		UOWHF_Result[6]:=UOWHF_Result[6] + 2040215044+UOWHF_Add_c;
   		UOWHF_Add_c.6:=UOWHF_Result[6].31;
   		UOWHF_Result[6].31:=0;
   	End_If;
   	If UOWHF_Msg[1].[29] Then
   		UOWHF_Result[0]:=UOWHF_Result[0] + 1358016563+UOWHF_Add_c;
   		UOWHF_Add_c.0:=UOWHF_Result[0].31;
   		UOWHF_Result[0].31:=0;
   		UOWHF_Result[1]:=UOWHF_Result[1] + 1270079032+UOWHF_Add_c;
   		UOWHF_Add_c.1:=UOWHF_Result[1].31;
   		UOWHF_Result[1].31:=0;
   		UOWHF_Result[2]:=UOWHF_Result[2] + 221615275+UOWHF_Add_c;
   		UOWHF_Add_c.2:=UOWHF_Result[2].31;
   		UOWHF_Result[2].31:=0;
   		UOWHF_Result[3]:=UOWHF_Result[3] + 122898292+UOWHF_Add_c;
   		UOWHF_Add_c.3:=UOWHF_Result[3].31;
   		UOWHF_Result[3].31:=0;
   		UOWHF_Result[4]:=UOWHF_Result[4] + 585819980+UOWHF_Add_c;
   		UOWHF_Add_c.4:=UOWHF_Result[4].31;
   		UOWHF_Result[4].31:=0;
   		UOWHF_Result[5]:=UOWHF_Result[5] + 51892856+UOWHF_Add_c;
   		UOWHF_Add_c.5:=UOWHF_Result[5].31;
   		UOWHF_Result[5].31:=0;
   		UOWHF_Result[6]:=UOWHF_Result[6] + 2033448244+UOWHF_Add_c;
   		UOWHF_Add_c.6:=UOWHF_Result[6].31;
   		UOWHF_Result[6].31:=0;
   	End_If;
   	If UOWHF_Msg[1].[30] Then
   		UOWHF_Result[0]:=UOWHF_Result[0] + 1133859205+UOWHF_Add_c;
   		UOWHF_Add_c.0:=UOWHF_Result[0].31;
   		UOWHF_Result[0].31:=0;
   		UOWHF_Result[1]:=UOWHF_Result[1] + 1230076861+UOWHF_Add_c;
   		UOWHF_Add_c.1:=UOWHF_Result[1].31;
   		UOWHF_Result[1].31:=0;
   		UOWHF_Result[2]:=UOWHF_Result[2] + 628374261+UOWHF_Add_c;
   		UOWHF_Add_c.2:=UOWHF_Result[2].31;
   		UOWHF_Result[2].31:=0;
   		UOWHF_Result[3]:=UOWHF_Result[3] + 528948219+UOWHF_Add_c;
   		UOWHF_Add_c.3:=UOWHF_Result[3].31;
   		UOWHF_Result[3].31:=0;
   		UOWHF_Result[4]:=UOWHF_Result[4] + 972509243+UOWHF_Add_c;
   		UOWHF_Add_c.4:=UOWHF_Result[4].31;
   		UOWHF_Result[4].31:=0;
   		UOWHF_Result[5]:=UOWHF_Result[5] + 2043873556+UOWHF_Add_c;
   		UOWHF_Add_c.5:=UOWHF_Result[5].31;
   		UOWHF_Result[5].31:=0;
   		UOWHF_Result[6]:=UOWHF_Result[6] + 1092533412+UOWHF_Add_c;
   		UOWHF_Add_c.6:=UOWHF_Result[6].31;
   		UOWHF_Result[6].31:=0;
   	End_If;
   	If UOWHF_Msg[1].[31] Then
   		UOWHF_Result[0]:=UOWHF_Result[0] + 1606040904+UOWHF_Add_c;
   		UOWHF_Add_c.0:=UOWHF_Result[0].31;
   		UOWHF_Result[0].31:=0;
   		UOWHF_Result[1]:=UOWHF_Result[1] + 1954021178+UOWHF_Add_c;
   		UOWHF_Add_c.1:=UOWHF_Result[1].31;
   		UOWHF_Result[1].31:=0;
   		UOWHF_Result[2]:=UOWHF_Result[2] + 2142650118+UOWHF_Add_c;
   		UOWHF_Add_c.2:=UOWHF_Result[2].31;
   		UOWHF_Result[2].31:=0;
   		UOWHF_Result[3]:=UOWHF_Result[3] + 608618905+UOWHF_Add_c;
   		UOWHF_Add_c.3:=UOWHF_Result[3].31;
   		UOWHF_Result[3].31:=0;
   		UOWHF_Result[4]:=UOWHF_Result[4] + 865412167+UOWHF_Add_c;
   		UOWHF_Add_c.4:=UOWHF_Result[4].31;
   		UOWHF_Result[4].31:=0;
   		UOWHF_Result[5]:=UOWHF_Result[5] + 181818924+UOWHF_Add_c;
   		UOWHF_Add_c.5:=UOWHF_Result[5].31;
   		UOWHF_Result[5].31:=0;
   		UOWHF_Result[6]:=UOWHF_Result[6] + 153939124+UOWHF_Add_c;
   		UOWHF_Add_c.6:=UOWHF_Result[6].31;
   		UOWHF_Result[6].31:=0;
   	End_If;
   	If UOWHF_Msg[2].[0] Then
   		UOWHF_Result[0]:=UOWHF_Result[0] + 162418271+UOWHF_Add_c;
   		UOWHF_Add_c.0:=UOWHF_Result[0].31;
   		UOWHF_Result[0].31:=0;
   		UOWHF_Result[1]:=UOWHF_Result[1] + 1022718455+UOWHF_Add_c;
   		UOWHF_Add_c.1:=UOWHF_Result[1].31;
   		UOWHF_Result[1].31:=0;
   		UOWHF_Result[2]:=UOWHF_Result[2] + 1321172784+UOWHF_Add_c;
   		UOWHF_Add_c.2:=UOWHF_Result[2].31;
   		UOWHF_Result[2].31:=0;
   		UOWHF_Result[3]:=UOWHF_Result[3] + 1943307377+UOWHF_Add_c;
   		UOWHF_Add_c.3:=UOWHF_Result[3].31;
   		UOWHF_Result[3].31:=0;
   		UOWHF_Result[4]:=UOWHF_Result[4] + 204552101+UOWHF_Add_c;
   		UOWHF_Add_c.4:=UOWHF_Result[4].31;
   		UOWHF_Result[4].31:=0;
   		UOWHF_Result[5]:=UOWHF_Result[5] + 935055409+UOWHF_Add_c;
   		UOWHF_Add_c.5:=UOWHF_Result[5].31;
   		UOWHF_Result[5].31:=0;
   		UOWHF_Result[6]:=UOWHF_Result[6] + 1030104506+UOWHF_Add_c;
   		UOWHF_Add_c.6:=UOWHF_Result[6].31;
   		UOWHF_Result[6].31:=0;
   	End_If;
   	If UOWHF_Msg[2].[1] Then
   		UOWHF_Result[0]:=UOWHF_Result[0] + 516643732+UOWHF_Add_c;
   		UOWHF_Add_c.0:=UOWHF_Result[0].31;
   		UOWHF_Result[0].31:=0;
   		UOWHF_Result[1]:=UOWHF_Result[1] + 1804822872+UOWHF_Add_c;
   		UOWHF_Add_c.1:=UOWHF_Result[1].31;
   		UOWHF_Result[1].31:=0;
   		UOWHF_Result[2]:=UOWHF_Result[2] + 310439864+UOWHF_Add_c;
   		UOWHF_Add_c.2:=UOWHF_Result[2].31;
   		UOWHF_Result[2].31:=0;
   		UOWHF_Result[3]:=UOWHF_Result[3] + 1619798537+UOWHF_Add_c;
   		UOWHF_Add_c.3:=UOWHF_Result[3].31;
   		UOWHF_Result[3].31:=0;
   		UOWHF_Result[4]:=UOWHF_Result[4] + 229400100+UOWHF_Add_c;
   		UOWHF_Add_c.4:=UOWHF_Result[4].31;
   		UOWHF_Result[4].31:=0;
   		UOWHF_Result[5]:=UOWHF_Result[5] + 2041405893+UOWHF_Add_c;
   		UOWHF_Add_c.5:=UOWHF_Result[5].31;
   		UOWHF_Result[5].31:=0;
   		UOWHF_Result[6]:=UOWHF_Result[6] + 658088462+UOWHF_Add_c;
   		UOWHF_Add_c.6:=UOWHF_Result[6].31;
   		UOWHF_Result[6].31:=0;
   	End_If;
   	If UOWHF_Msg[2].[2] Then
   		UOWHF_Result[0]:=UOWHF_Result[0] + 163619853+UOWHF_Add_c;
   		UOWHF_Add_c.0:=UOWHF_Result[0].31;
   		UOWHF_Result[0].31:=0;
   		UOWHF_Result[1]:=UOWHF_Result[1] + 1055853189+UOWHF_Add_c;
   		UOWHF_Add_c.1:=UOWHF_Result[1].31;
   		UOWHF_Result[1].31:=0;
   		UOWHF_Result[2]:=UOWHF_Result[2] + 1496964915+UOWHF_Add_c;
   		UOWHF_Add_c.2:=UOWHF_Result[2].31;
   		UOWHF_Result[2].31:=0;
   		UOWHF_Result[3]:=UOWHF_Result[3] + 1875623055+UOWHF_Add_c;
   		UOWHF_Add_c.3:=UOWHF_Result[3].31;
   		UOWHF_Result[3].31:=0;
   		UOWHF_Result[4]:=UOWHF_Result[4] + 1628553455+UOWHF_Add_c;
   		UOWHF_Add_c.4:=UOWHF_Result[4].31;
   		UOWHF_Result[4].31:=0;
   		UOWHF_Result[5]:=UOWHF_Result[5] + 2128870259+UOWHF_Add_c;
   		UOWHF_Add_c.5:=UOWHF_Result[5].31;
   		UOWHF_Result[5].31:=0;
   		UOWHF_Result[6]:=UOWHF_Result[6] + 1009565693+UOWHF_Add_c;
   		UOWHF_Add_c.6:=UOWHF_Result[6].31;
   		UOWHF_Result[6].31:=0;
   	End_If;
   	If UOWHF_Msg[2].[3] Then
   		UOWHF_Result[0]:=UOWHF_Result[0] + 22660734+UOWHF_Add_c;
   		UOWHF_Add_c.0:=UOWHF_Result[0].31;
   		UOWHF_Result[0].31:=0;
   		UOWHF_Result[1]:=UOWHF_Result[1] + 2045680470+UOWHF_Add_c;
   		UOWHF_Add_c.1:=UOWHF_Result[1].31;
   		UOWHF_Result[1].31:=0;
   		UOWHF_Result[2]:=UOWHF_Result[2] + 161249708+UOWHF_Add_c;
   		UOWHF_Add_c.2:=UOWHF_Result[2].31;
   		UOWHF_Result[2].31:=0;
   		UOWHF_Result[3]:=UOWHF_Result[3] + 1005315890+UOWHF_Add_c;
   		UOWHF_Add_c.3:=UOWHF_Result[3].31;
   		UOWHF_Result[3].31:=0;
   		UOWHF_Result[4]:=UOWHF_Result[4] + 1356423176+UOWHF_Add_c;
   		UOWHF_Add_c.4:=UOWHF_Result[4].31;
   		UOWHF_Result[4].31:=0;
   		UOWHF_Result[5]:=UOWHF_Result[5] + 1710579281+UOWHF_Add_c;
   		UOWHF_Add_c.5:=UOWHF_Result[5].31;
   		UOWHF_Result[5].31:=0;
   		UOWHF_Result[6]:=UOWHF_Result[6] + 1524950966+UOWHF_Add_c;
   		UOWHF_Add_c.6:=UOWHF_Result[6].31;
   		UOWHF_Result[6].31:=0;
   	End_If;
   	If UOWHF_Msg[2].[4] Then
   		UOWHF_Result[0]:=UOWHF_Result[0] + 1634981150+UOWHF_Add_c;
   		UOWHF_Add_c.0:=UOWHF_Result[0].31;
   		UOWHF_Result[0].31:=0;
   		UOWHF_Result[1]:=UOWHF_Result[1] + 1394453812+UOWHF_Add_c;
   		UOWHF_Add_c.1:=UOWHF_Result[1].31;
   		UOWHF_Result[1].31:=0;
   		UOWHF_Result[2]:=UOWHF_Result[2] + 287411036+UOWHF_Add_c;
   		UOWHF_Add_c.2:=UOWHF_Result[2].31;
   		UOWHF_Result[2].31:=0;
   		UOWHF_Result[3]:=UOWHF_Result[3] + 1956843077+UOWHF_Add_c;
   		UOWHF_Add_c.3:=UOWHF_Result[3].31;